HMI tags "MixingHead"
   "DB611_Hydraulic_State_Read" : Bool = PLC DB611_Hydraulic_State.Read AT %DB611.DBX8.0, 1 s
   "DB611_Hydraulic_State_Write" : Bool = PLC DB14_TP_Shortcuts.TP_Shortcuts.PageNo.7 AT %DB611.DBX8.1, 1 s
   "DB721_MH_Hydraulic_MH_Hyd{0}_Hyd_CP_Time" : S5Time = PLC DB14_TP_Shortcuts.TP_Shortcuts.PageNo.3 AT %DB721.DBW18, 1 s
      on ChangeValue: SetBit("DB611_Hydraulic_State_Write")
   "DB721_MH_Hydraulic_MH_Hyd{0}_Hyd_P_Startup" : S5Time = PLC DB14_TP_Shortcuts.TP_Shortcuts.PageNo.2 AT %DB721.DBW14, 1 s
      on ChangeValue: SetBit("DB611_Hydraulic_State_Write")
   "DB721_MH_Hydraulic_MH_Hyd{0}_Hyd_P_Supervision" : S5Time = PLC DB14_TP_Shortcuts.TP_Shortcuts.PageNo.4 AT %DB721.DBW16, 1 s
      on ChangeValue: SetBit("DB611_Hydraulic_State_Write")
   "DB721_MH_Hydraulic_MH_Hyd{0}_Hyd_PressureSwitch" : S5Time = PLC DB14_TP_Shortcuts.TP_Shortcuts.PageNo.5 AT %DB721.DBW20, 1 s
      on ChangeValue: SetBit("DB611_Hydraulic_State_Write")
   "DB721_MH_Hydraulic_MH_Hyd{0}_Hyd_SwitchOFFDelay" : S5Time = PLC DB14_TP_Shortcuts.TP_Shortcuts.PageNo.6 AT %DB721.DBW22, 1 s
      on ChangeValue: SetBit("DB611_Hydraulic_State_Write")
   "DB721_MH_Hydraulic_Option{0}_With2PSwitch" : Bool = PLC DB721_MH_Hydraulic.Option[0].With2PSwitch AT %DB721.DBX6.0, 1 s
   "MixingHead Options" : Int, internal
   "DB704_MH_Value_Read" : Bool = PLC DB704_MH_Value.Read AT %DB704.DBX4.0, 1 s
   "DB614_MH_State_Read" : Bool = PLC DB614_MH_State.Read AT %DB614.DBX8.0, 1 s
   "DB614_MH_State_Write" : Bool = PLC DB614_MH_State.Write AT %DB614.DBX8.1, 1 s
   "DB614_MH_State_MH_Status{0}_QPB_Values_selected" : Bool = PLC DB614_MH_State.MH_Status[0].QPB_Values_selected AT %DB614.DBX3920.2, 1 s
   "DB704_MH_Value_MH_Inerting{0}_Purge_time" : S5Time = PLC DB704_MH_Value.MH_Inerting[0].Purge_time AT %DB704.DBW4568, 1 s
      on ChangeValue: SetBit("DB704_MH_Value_Write")
   "DB704_MH_Value_MH_Inerting{0}_Purge_after_Shot" : S5Time = PLC DB704_MH_Value.MH_Inerting[0].Purge_after_Shot AT %DB704.DBW4570, 1 s
      on ChangeValue: SetBit("DB704_MH_Value_Write")
   "DB704_MH_Value_Mixinghead{0}_MH_Connection{1}_Flow_red_Circ" : Real = PLC DB704_MH_Value.Mixinghead[0].MH_Connection[1].Flow_red_Circ AT %DB704.DBD74, 1 s
      on ChangeValue: SetBit("DB704_MH_Value_Write")
   "DB704_MH_Value_Mixinghead{0}_MH_Connection{1}_Flow_HP_Circ" : Real = PLC DB704_MH_Value.Mixinghead[0].MH_Connection[1].Flow_HP_Circ AT %DB704.DBD70, 1 s
      on ChangeValue: SetBit("DB704_MH_Value_Write")
   "DB704_MH_Value_Mixinghead{0}_MH_Connection{1}_Flow_LP_Circ" : Real = PLC DB704_MH_Value.Mixinghead[0].MH_Connection[1].Flow_LP_Circ AT %DB704.DBD78, 1 s
      on ChangeValue: SetBit("DB704_MH_Value_Write")
   "DB704_MH_Value_Mixinghead{0}_MH_Connection{2}_Flow_HP_Circ" : Real = PLC DB704_MH_Value.Mixinghead[0].MH_Connection[2].Flow_HP_Circ AT %DB704.DBD104, 1 s
      on ChangeValue: SetBit("DB704_MH_Value_Write")
   "DB704_MH_Value_Mixinghead{0}_MH_Connection{2}_Flow_red_Circ" : Real = PLC DB704_MH_Value.Mixinghead[0].MH_Connection[2].Flow_red_Circ AT %DB704.DBD108, 1 s
      on ChangeValue: SetBit("DB704_MH_Value_Write")
   "DB704_MH_Value_Mixinghead{0}_MH_Connection{2}_Flow_LP_Circ" : Real = PLC DB704_MH_Value.Mixinghead[0].MH_Connection[2].Flow_LP_Circ AT %DB704.DBD112, 1 s
      on ChangeValue: SetBit("DB704_MH_Value_Write")
   "DB704_MH_Value_Mixinghead{0}_MH_Connection{1}_FlowQPB" : Real = PLC DB704_MH_Value.Mixinghead[0].MH_Connection[1].FlowQPB AT %DB704.DBD90, 1 s
      on ChangeValue: SetBit("DB704_MH_Value_Write")
   "DB704_MH_Value_Mixinghead{0}_MH_Connection{1}_HP_CircOverNozzle" : Bool = PLC DB704_MH_Value.Mixinghead[0].MH_Connection[1].HP_CircOverNozzle AT %DB704.DBX98.0, 1 s
      on ChangeValue: SetBit("DB614_MH_State_Write")
   "DB704_MH_Value_Mixinghead{0}_MH_Connection{1}_Red_CircOverNozzle" : Bool = PLC DB704_MH_Value.Mixinghead[0].MH_Connection[1].Red_CircOverNozzle AT %DB704.DBX98.1, 1 s
      on ChangeValue: SetBit("DB614_MH_State_Write")
   "DB704_MH_Value_Mixinghead{0}_MH_Connection{1}_LP_CircOverNozzle" : Bool = PLC DB704_MH_Value.Mixinghead[0].MH_Connection[1].LP_CircOverNozzle AT %DB704.DBX98.2, 1 s
      on ChangeValue: SetBit("DB614_MH_State_Write")
   "DB704_MH_Value_Mixinghead{0}_MH_Connection{2}_HP_CircOverNozzle" : Bool = PLC DB704_MH_Value.Mixinghead[0].MH_Connection[2].HP_CircOverNozzle AT %DB704.DBX132.0, 1 s
      on ChangeValue: SetBit("DB614_MH_State_Write")
   "DB704_MH_Value_Mixinghead{0}_MH_Connection{2}_Red_CircOverNozzle" : Bool = PLC DB704_MH_Value.Mixinghead[0].MH_Connection[2].Red_CircOverNozzle AT %DB704.DBX132.1, 1 s
      on ChangeValue: SetBit("DB614_MH_State_Write")
   "DB704_MH_Value_Mixinghead{0}_MH_Connection{2}_LP_CircOverNozzle" : Bool = PLC DB704_MH_Value.Mixinghead[0].MH_Connection[2].LP_CircOverNozzle AT %DB704.DBX132.2, 1 s
      on ChangeValue: SetBit("DB614_MH_State_Write")
   "MH_Control_Visibility" : Int AT %DB1.DBX0.0
   "DB704_MH_Value_Mixinghead{0}_MH_Connection{2}_FlowQPB" : Real = PLC DB704_MH_Value.Mixinghead[0].MH_Connection[2].FlowQPB AT %DB704.DBD124, 1 s
      on ChangeValue: SetBit("DB704_MH_Value_Write")
   "DB704_MH_Value_Mixinghead{0}_MH_Connection{2}_PressureQPB" : Real = PLC DB704_MH_Value.Mixinghead[0].MH_Connection[2].PressureQPB AT %DB704.DBD128, 1 s
      on ChangeValue: SetBit("DB704_MH_Value_Write")
   "DB704_MH_Value_Mixinghead{0}_MH_Connection{1}_PressureQPB" : Real = PLC DB704_MH_Value.Mixinghead[0].MH_Connection[1].PressureQPB AT %DB704.DBD94, 1 s
      on ChangeValue: SetBit("DB704_MH_Value_Write")
   "DB704_MH_Value_Mixinghead{0}_Cleaning_Piston_RestTimeBack" : S5Time = PLC DB704_MH_Value.Mixinghead[0].Cleaning_Piston.RestTimeBack AT %DB704.DBW44, 1 s
      on ChangeValue: SetBit("DB704_MH_Value_Write")
   "DB704_MH_Value_Mixinghead{0}_Cleaning_Piston_RestTimeFront" : S5Time = PLC DB704_MH_Value.Mixinghead[0].Cleaning_Piston.RestTimeFront AT %DB704.DBW46, 1 s
      on ChangeValue: SetBit("DB704_MH_Value_Write")
   "DB704_MH_Value_Mixinghead{0}_Cleaning_Piston_RestTimeFrontManual" : S5Time = PLC DB704_MH_Value.Mixinghead[0].Cleaning_Piston.RestTimeFrontManual AT %DB704.DBW48, 1 s
      on ChangeValue: SetBit("DB704_MH_Value_Write")
   "DB704_MH_Value_Write" : Bool = PLC DB704_MH_Value.Write AT %DB704.DBX4.1, 1 s
   "DB704_MH_Value_MH_Inerting{0}_Max_Inerting_Time" : S5Time = PLC DB704_MH_Value.MH_Inerting[0].Max_Inerting_Time AT %DB704.DBW4560, 1 s
      on ChangeValue: SetBit("DB704_MH_Value_Write")
   "DB704_MH_Value_MH_Inerting{0}_Ready_Time_after_Inert" : S5Time = PLC DB704_MH_Value.MH_Inerting[0].Ready_Time_after_Inert AT %DB704.DBW4562, 1 s
      on ChangeValue: SetBit("DB704_MH_Value_Write")
   "DB704_MH_Value_MH_Inerting{0}_Foam_density" : DInt = PLC DB704_MH_Value.MH_Inerting[0].Foam_density AT %DB704.DBD4538, 1 s
      on ChangeValue: SetBit("DB704_MH_Value_Write")
   "DB704_MH_Value_MH_Inerting{0}_Inerting_factor" : Real = PLC DB704_MH_Value.MH_Inerting[0].Inerting_factor AT %DB704.DBD4542, 1 s
      on ChangeValue: SetBit("DB704_MH_Value_Write")
   "DB704_MH_Value_MH_Inerting{0}_Start_Offset" : Real = PLC DB704_MH_Value.MH_Inerting[0].Start_Offset AT %DB704.DBD4546, 1 s
      on ChangeValue: SetBit("DB704_MH_Value_Write")
   "DB704_MH_Value_MH_Inerting{0}_Leakage_Value" : Real = PLC DB704_MH_Value.MH_Inerting[0].Leakage_Value AT %DB704.DBD4550, 1 s
      on ChangeValue: SetBit("DB704_MH_Value_Write")
   "DB704_MH_Value_Mixinghead{0}_AmountComponent" : Byte = PLC DB704_MH_Value.Mixinghead[0].AmountComponent AT %DB704.DBB6, 1 s
      on ChangeValue: SetBit("DB704_MH_Value_Write")
   "DB704_MH_Value_Mixinghead{0}_MachineNumber" : Byte = PLC DB704_MH_Value.Mixinghead[0].MachineNumber AT %DB704.DBB7, 1 s
      on ChangeValue: SetBit("DB704_MH_Value_Write")
   "DB704_MH_Value_Mixinghead{0}_MH_Active" : Bool = PLC DB704_MH_Value.Mixinghead[0].MH_Active AT %DB704.DBX9.0, 1 s
      on ChangeValue: SetBit("DB614_MH_State_Write")
   "DB704_MH_Value_Mixinghead{0}_With99program" : Bool = PLC DB704_MH_Value.Mixinghead[0].With99program AT %DB704.DBX10.2, 1 s
      on ChangeValue: SetBit("DB704_MH_Value_Write")
   "DB704_MH_Value_Mixinghead{0}_WithHeating" : Bool = PLC DB704_MH_Value.Mixinghead[0].WithHeating AT %DB704.DBX9.6, 1 s
      on ChangeValue: SetBit("DB704_MH_Value_Write")
   "DB704_MH_Value_Mixinghead{0}_WithInerting" : Bool = PLC DB704_MH_Value.Mixinghead[0].WithInerting AT %DB704.DBX9.5, 1 s
      on ChangeValue: SetBit("DB704_MH_Value_Write")
   "DB704_MH_Value_Mixinghead{0}_WithInterface" : Bool = PLC DB704_MH_Value.Mixinghead[0].WithInterface AT %DB704.DBX9.4, 1 s
      on ChangeValue: SetBit("DB704_MH_Value_Write")
   "DB704_MH_Value_Mixinghead{0}_WithNozzleControl" : Bool = PLC DB704_MH_Value.Mixinghead[0].WithNozzleControl AT %DB704.DBX9.2, 1 s
      on ChangeValue: SetBit("DB704_MH_Value_Write")
   "DB704_MH_Value_Mixinghead{0}_WithCleaningPiston" : Bool = PLC DB704_MH_Value.Mixinghead[0].WithCleaningPiston AT %DB704.DBX9.1, 1 s
      on ChangeValue: SetBit("DB704_MH_Value_Write")
   "DB704_MH_Value_Mixinghead{0}_WithLPCirculation" : Bool = PLC DB704_MH_Value.Mixinghead[0].WithLPCirculation AT %DB704.DBX9.3, 1 s
      on ChangeValue: SetBit("DB704_MH_Value_Write")
   "DB704_MH_Value_Mixinghead{0}_pRrgNumberManual" : Byte = PLC DB704_MH_Value.Mixinghead[0].pRrgNumberManual AT %DB704.DBB8, 1 s
      on ChangeValue: SetBit("DB704_MH_Value_Write")
   "DB704_MH_Value_Mixinghead{0}_Openingtime" : Real = PLC DB704_MH_Value.Mixinghead[0].Openingtime AT %DB704.DBD14, 1 s
      on ChangeValue: SetBit("DB704_MH_Value_Write")
   "DB704_MH_Value_Mixinghead{0}_Closingtime" : Real = PLC DB704_MH_Value.Mixinghead[0].Closingtime AT %DB704.DBD18, 1 s
      on ChangeValue: SetBit("DB704_MH_Value_Write")
   "DB604_PV_Mixinghead_Mixinghead{0}_Temperature_Connection{1}_PV_ActV_Value" : Real = PLC DB604_PV_Mixinghead.Mixinghead[0].Temperature_Connection[1].PV_ActV.Value AT %DB604.DBD314, 1 s
      on ChangeValue: SetBit("DB704_MH_Value_Write")
   "DB604_PV_Mixinghead_Mixinghead{0}_Temperature_Connection{1}_PV_SetV_Value" : Real = PLC DB604_PV_Mixinghead.Mixinghead[0].Temperature_Connection[1].PV_SetV.Value AT %DB604.DBD294, 1 s
      on ChangeValue: SetBit("DB704_MH_Value_Write")
   "DB604_PV_Mixinghead_Mixinghead{0}_Temperature_Connection{1}_PV_SetV_WarningLowerLimit" : Real = PLC DB604_PV_Mixinghead.Mixinghead[0].Temperature_Connection[1].PV_SetV.WarningLowerLimit AT %DB604.DBD298, 1 s
      on ChangeValue: SetBit("DB704_MH_Value_Write")
   "DB604_PV_Mixinghead_Mixinghead{0}_Temperature_Connection{1}_PV_SetV_WarningUpperLimit" : Real = PLC DB604_PV_Mixinghead.Mixinghead[0].Temperature_Connection[1].PV_SetV.WarningUpperLimit AT %DB604.DBD302, 1 s
      on ChangeValue: SetBit("DB704_MH_Value_Write")
   "DB604_PV_Mixinghead_Mixinghead{0}_Temperature_Connection{1}_PV_SetV_AlarmLowerLimit" : Real = PLC DB604_PV_Mixinghead.Mixinghead[0].Temperature_Connection[1].PV_SetV.AlarmLowerLimit AT %DB604.DBD306, 1 s
      on ChangeValue: SetBit("DB704_MH_Value_Write")
   "DB604_PV_Mixinghead_Mixinghead{0}_Temperature_Connection{1}_PV_SetV_AlarmUpperLimit" : Real = PLC DB604_PV_Mixinghead.Mixinghead[0].Temperature_Connection[1].PV_SetV.AlarmUpperLimit AT %DB604.DBD310, 1 s
      on ChangeValue: SetBit("DB704_MH_Value_Write")
   "DB604_PV_Mixinghead_Mixinghead{0}_Pressure_Connection{1}_PV_SetV_Value" : Real = PLC DB604_PV_Mixinghead.Mixinghead[0].Pressure_Connection[1].PV_SetV.Value AT %DB604.DBD6, 1 s
      on ChangeValue: SetBit("DB704_MH_Value_Write")
   "DB604_PV_Mixinghead_Mixinghead{0}_Pressure_Connection{1}_PV_SetV_WarningLowerLimit" : Real = PLC DB604_PV_Mixinghead.Mixinghead[0].Pressure_Connection[1].PV_SetV.WarningLowerLimit AT %DB604.DBD10, 1 s
      on ChangeValue: SetBit("DB704_MH_Value_Write")
   "DB604_PV_Mixinghead_Mixinghead{0}_Pressure_Connection{1}_PV_SetV_WarningUpperLimit" : Real = PLC DB604_PV_Mixinghead.Mixinghead[0].Pressure_Connection[1].PV_SetV.WarningUpperLimit AT %DB604.DBD14, 1 s
      on ChangeValue: SetBit("DB704_MH_Value_Write")
   "DB604_PV_Mixinghead_Mixinghead{0}_Pressure_Connection{1}_PV_SetV_AlarmLowerLimit" : Real = PLC DB604_PV_Mixinghead.Mixinghead[0].Pressure_Connection[1].PV_SetV.AlarmLowerLimit AT %DB604.DBD18, 1 s
      on ChangeValue: SetBit("DB704_MH_Value_Write")
   "DB604_PV_Mixinghead_Mixinghead{0}_Pressure_Connection{1}_PV_SetV_AlarmUpperLimit" : Real = PLC DB604_PV_Mixinghead.Mixinghead[0].Pressure_Connection[1].PV_SetV.AlarmUpperLimit AT %DB604.DBD22, 1 s
      on ChangeValue: SetBit("DB704_MH_Value_Write")
   "DB604_PV_Mixinghead_Mixinghead{0}_Pressure_Connection{1}_PV_ActV_Value" : Real = PLC DB604_PV_Mixinghead.Mixinghead[0].Pressure_Connection[1].PV_ActV.Value AT %DB604.DBD26, 1 s
      on ChangeValue: SetBit("DB704_MH_Value_Write")
   "DB604_PV_Mixinghead_Mixinghead{0}_Pressure_Connection{2}_PV_SetV_Value" : Real = PLC DB604_PV_Mixinghead.Mixinghead[0].Pressure_Connection[2].PV_SetV.Value AT %DB604.DBD54, 1 s
      on ChangeValue: SetBit("DB704_MH_Value_Write")
   "DB604_PV_Mixinghead_Mixinghead{0}_Pressure_Connection{2}_PV_SetV_WarningLowerLimit" : Real = PLC DB604_PV_Mixinghead.Mixinghead[0].Pressure_Connection[2].PV_SetV.WarningLowerLimit AT %DB604.DBD58, 1 s
      on ChangeValue: SetBit("DB704_MH_Value_Write")
   "DB604_PV_Mixinghead_Mixinghead{0}_Pressure_Connection{2}_PV_SetV_WarningUpperLimit" : Real = PLC DB604_PV_Mixinghead.Mixinghead[0].Pressure_Connection[2].PV_SetV.WarningUpperLimit AT %DB604.DBD62, 1 s
      on ChangeValue: SetBit("DB704_MH_Value_Write")
   "DB604_PV_Mixinghead_Mixinghead{0}_Pressure_Connection{2}_PV_SetV_AlarmLowerLimit" : Real = PLC DB604_PV_Mixinghead.Mixinghead[0].Pressure_Connection[2].PV_SetV.AlarmLowerLimit AT %DB604.DBD66, 1 s
      on ChangeValue: SetBit("DB704_MH_Value_Write")
   "DB604_PV_Mixinghead_Mixinghead{0}_Pressure_Connection{2}_PV_SetV_AlarmUpperLimit" : Real = PLC DB604_PV_Mixinghead.Mixinghead[0].Pressure_Connection[2].PV_SetV.AlarmUpperLimit AT %DB604.DBD70, 1 s
      on ChangeValue: SetBit("DB704_MH_Value_Write")
   "DB604_PV_Mixinghead_Mixinghead{0}_Pressure_Connection{2}_PV_ActV_Value" : Real = PLC DB604_PV_Mixinghead.Mixinghead[0].Pressure_Connection[2].PV_ActV.Value AT %DB604.DBD74, 1 s
      on ChangeValue: SetBit("DB704_MH_Value_Write")
   "DB604_PV_Mixinghead_Mixinghead{0}_Temperature_Connection{2}_PV_SetV_Value" : Real = PLC DB604_PV_Mixinghead.Mixinghead[0].Temperature_Connection[2].PV_SetV.Value AT %DB604.DBD342, 1 s
      on ChangeValue: SetBit("DB704_MH_Value_Write")
   "DB604_PV_Mixinghead_Mixinghead{0}_Temperature_Connection{2}_PV_SetV_WarningLowerLimit" : Real = PLC DB604_PV_Mixinghead.Mixinghead[0].Temperature_Connection[2].PV_SetV.WarningLowerLimit AT %DB604.DBD346, 1 s
      on ChangeValue: SetBit("DB704_MH_Value_Write")
   "DB604_PV_Mixinghead_Mixinghead{0}_Temperature_Connection{2}_PV_SetV_WarningUpperLimit" : Real = PLC DB604_PV_Mixinghead.Mixinghead[0].Temperature_Connection[2].PV_SetV.WarningUpperLimit AT %DB604.DBD350, 1 s
      on ChangeValue: SetBit("DB704_MH_Value_Write")
   "DB604_PV_Mixinghead_Mixinghead{0}_Temperature_Connection{2}_PV_SetV_AlarmLowerLimit" : Real = PLC DB604_PV_Mixinghead.Mixinghead[0].Temperature_Connection[2].PV_SetV.AlarmLowerLimit AT %DB604.DBD354, 1 s
      on ChangeValue: SetBit("DB704_MH_Value_Write")
   "DB604_PV_Mixinghead_Mixinghead{0}_Temperature_Connection{2}_PV_SetV_AlarmUpperLimit" : Real = PLC DB604_PV_Mixinghead.Mixinghead[0].Temperature_Connection[2].PV_SetV.AlarmUpperLimit AT %DB604.DBD358, 1 s
      on ChangeValue: SetBit("DB704_MH_Value_Write")
   "DB604_PV_Mixinghead_Mixinghead{0}_Temperature_Connection{2}_PV_ActV_Value" : Real = PLC DB604_PV_Mixinghead.Mixinghead[0].Temperature_Connection[2].PV_ActV.Value AT %DB604.DBD362, 1 s
      on ChangeValue: SetBit("DB704_MH_Value_Write")
   "DB704_MH_Value_Mixinghead{0}_Cleaning_Piston_CP_withInterval" : Bool = PLC DB704_MH_Value.Mixinghead[0].Cleaning_Piston.CP_withInterval AT %DB704.DBX56.1, 1 s
      on ChangeValue: SetBit("DB704_MH_Value_Write")
   "DB704_MH_Value_Mixinghead{0}_Cleaning_Piston_ContrCleaningPiston" : Bool = PLC DB704_MH_Value.Mixinghead[0].Cleaning_Piston.ContrCleaningPiston AT %DB704.DBX56.3, 1 s
      on ChangeValue: SetBit("DB704_MH_Value_Write")
   "DB611_Hydraulic_State_MH_Hydraulic{0}_HourCounter" : DInt = PLC DB611_Hydraulic_State.MH_Hydraulic[0].HourCounter AT %DB611.DBD14, 1 s
   "DB614_MH_State_ReadDeviceNo" : Int = PLC DB614_MH_State.ReadDeviceNo AT %DB614.DBW0, 1 s
   "DB704_MH_Value_Mixinghead{0}_WithMHVenting" : Bool = PLC DB704_MH_Value.Mixinghead[0].WithMHVenting AT %DB704.DBX9.7, 1 s
      on ChangeValue: SetBit("DB704_MH_Value_Write")
   "DB614_MH_State_MH_Status{0}_Switch_HP_ON_OFF" : Bool = PLC DB614_MH_State.MH_Status[0].Switch_HP_ON_OFF AT %DB614.DBX3920.5, 1 s
      on ChangeValue: SetBit("DB614_MH_State_Write")
   "DB614_MH_State_MH_Status{0}_Switch_Service_ON_OFF" : Bool = PLC DB614_MH_State.MH_Status[0].Switch_Service_ON_OFF AT %DB614.DBX3920.6, 1 s
      on ChangeValue: SetBit("DB614_MH_State_Write")
   "DB704_MH_Value_Mixinghead{0}_MH_Connection{3}_Flow_HP_Circ" : Real = PLC DB704_MH_Value.Mixinghead[0].MH_Connection[3].Flow_HP_Circ AT %DB704.DBD138, 1 s
   "DB704_MH_Value_Mixinghead{0}_MH_Connection{3}_Flow_red_Circ" : Real = PLC DB704_MH_Value.Mixinghead[0].MH_Connection[3].Flow_red_Circ AT %DB704.DBD142, 1 s
   "DB704_MH_Value_Mixinghead{0}_MH_Connection{3}_Flow_LP_Circ" : Real = PLC DB704_MH_Value.Mixinghead[0].MH_Connection[3].Flow_LP_Circ AT %DB704.DBD146, 1 s
   "DB704_MH_Value_Mixinghead{0}_MH_Connection{3}_HP_CircOverNozzle" : Bool = PLC DB704_MH_Value.Mixinghead[0].MH_Connection[3].HP_CircOverNozzle AT %DB704.DBX166.0, 1 s
   "DB704_MH_Value_Mixinghead{0}_MH_Connection{3}_Red_CircOverNozzle" : Bool = PLC DB704_MH_Value.Mixinghead[0].MH_Connection[3].Red_CircOverNozzle AT %DB704.DBX166.1, 1 s
   "DB704_MH_Value_Mixinghead{0}_MH_Connection{3}_LP_CircOverNozzle" : Bool = PLC DB704_MH_Value.Mixinghead[0].MH_Connection[3].LP_CircOverNozzle AT %DB704.DBX166.2, 1 s
   "DB704_MH_Value_Mixinghead{0}_MH_Connection{4}_Flow_HP_Circ" : Real = PLC DB704_MH_Value.Mixinghead[0].MH_Connection[4].Flow_HP_Circ AT %DB704.DBD172, 1 s
   "DB704_MH_Value_Mixinghead{0}_MH_Connection{4}_Flow_red_Circ" : Real = PLC DB704_MH_Value.Mixinghead[0].MH_Connection[4].Flow_red_Circ AT %DB704.DBD176, 1 s
   "DB704_MH_Value_Mixinghead{0}_MH_Connection{4}_Flow_LP_Circ" : Real = PLC DB704_MH_Value.Mixinghead[0].MH_Connection[4].Flow_LP_Circ AT %DB704.DBD180, 1 s
   "DB704_MH_Value_Mixinghead{0}_MH_Connection{4}_HP_CircOverNozzle" : Bool = PLC DB704_MH_Value.Mixinghead[0].MH_Connection[4].HP_CircOverNozzle AT %DB704.DBX200.0, 1 s
   "DB704_MH_Value_Mixinghead{0}_MH_Connection{4}_Red_CircOverNozzle" : Bool = PLC DB702_Tank_Value.Tank[0].With_Drain AT %DB704.DBX200.1, 1 s
   "DB704_MH_Value_Mixinghead{0}_MH_Connection{4}_LP_CircOverNozzle" : Bool = PLC DB704_MH_Value.Mixinghead[0].MH_Connection[4].LP_CircOverNozzle AT %DB704.DBX200.2, 1 s
   "DB704_MH_Value_Mixinghead{0}_MH_Connection{5}_Flow_HP_Circ" : Real = PLC DB704_MH_Value.Mixinghead[0].MH_Connection[5].Flow_HP_Circ AT %DB704.DBD206, 1 s
   "DB704_MH_Value_Mixinghead{0}_MH_Connection{5}_Flow_red_Circ" : Real = PLC DB704_MH_Value.Mixinghead[0].MH_Connection[5].Flow_red_Circ AT %DB704.DBD210, 1 s
   "DB704_MH_Value_Mixinghead{0}_MH_Connection{5}_Flow_LP_Circ" : Real = PLC DB704_MH_Value.Mixinghead[0].MH_Connection[5].Flow_LP_Circ AT %DB704.DBD214, 1 s
   "DB704_MH_Value_Mixinghead{0}_MH_Connection{5}_HP_CircOverNozzle" : Bool = PLC DB704_MH_Value.Mixinghead[0].MH_Connection[5].HP_CircOverNozzle AT %DB704.DBX234.0, 1 s
   "DB704_MH_Value_Mixinghead{0}_MH_Connection{5}_Red_CircOverNozzle" : Bool = PLC DB704_MH_Value.Mixinghead[0].MH_Connection[5].Red_CircOverNozzle AT %DB704.DBX234.1, 1 s
   "DB704_MH_Value_Mixinghead{0}_MH_Connection{5}_LP_CircOverNozzle" : Bool = PLC DB704_MH_Value.Mixinghead[0].MH_Connection[5].LP_CircOverNozzle AT %DB704.DBX234.2, 1 s
   "DB704_MH_Value_Mixinghead{0}_MH_Connection{6}_Flow_HP_Circ" : Real = PLC DB704_MH_Value.Mixinghead[0].MH_Connection[6].Flow_HP_Circ AT %DB704.DBD240, 1 s
   "DB704_MH_Value_Mixinghead{0}_MH_Connection{6}_Flow_red_Circ" : Real = PLC DB704_MH_Value.Mixinghead[0].MH_Connection[6].Flow_red_Circ AT %DB704.DBD244, 1 s
   "DB704_MH_Value_Mixinghead{0}_MH_Connection{6}_Flow_LP_Circ" : Real = PLC DB704_MH_Value.Mixinghead[0].MH_Connection[6].Flow_LP_Circ AT %DB704.DBD248, 1 s
   "DB704_MH_Value_Mixinghead{0}_MH_Connection{6}_HP_CircOverNozzle" : Bool = PLC DB704_MH_Value.Mixinghead[0].MH_Connection[6].HP_CircOverNozzle AT %DB704.DBX268.0, 1 s
   "DB704_MH_Value_Mixinghead{0}_MH_Connection{6}_Red_CircOverNozzle" : Bool = PLC DB704_MH_Value.Mixinghead[0].MH_Connection[6].Red_CircOverNozzle AT %DB704.DBX268.1, 1 s
   "DB704_MH_Value_Mixinghead{0}_MH_Connection{6}_LP_CircOverNozzle" : Bool = PLC DB704_MH_Value.Mixinghead[0].MH_Connection[6].LP_CircOverNozzle AT %DB704.DBX268.2, 1 s
   "DB704_MH_Value_Mixinghead{0}_MH_Connection{3}_FlowQPB" : Real = PLC DB704_MH_Value.Mixinghead[0].MH_Connection[3].FlowQPB AT %DB704.DBD158, 1 s
   "DB704_MH_Value_Mixinghead{0}_MH_Connection{3}_PressureQPB" : Real = PLC DB704_MH_Value.Mixinghead[0].MH_Connection[3].PressureQPB AT %DB704.DBD162, 1 s
   "DB704_MH_Value_Mixinghead{0}_MH_Connection{4}_FlowQPB" : Real = PLC DB704_MH_Value.Mixinghead[0].MH_Connection[4].FlowQPB AT %DB704.DBD192, 1 s
   "DB704_MH_Value_Mixinghead{0}_MH_Connection{4}_PressureQPB" : Real = PLC DB704_MH_Value.Mixinghead[0].MH_Connection[4].PressureQPB AT %DB704.DBD196, 1 s
   "DB704_MH_Value_Mixinghead{0}_MH_Connection{5}_FlowQPB" : Real = PLC DB704_MH_Value.Mixinghead[0].MH_Connection[5].FlowQPB AT %DB704.DBD226, 1 s
   "DB704_MH_Value_Mixinghead{0}_MH_Connection{5}_PressureQPB" : Real = PLC DB704_MH_Value.Mixinghead[0].MH_Connection[5].PressureQPB AT %DB704.DBD230, 1 s
   "DB704_MH_Value_Mixinghead{0}_MH_Connection{6}_FlowQPB" : Real = PLC DB704_MH_Value.Mixinghead[0].MH_Connection[6].FlowQPB AT %DB704.DBD260, 1 s
   "DB704_MH_Value_Mixinghead{0}_MH_Connection{6}_PressureQPB" : Real = PLC DB704_MH_Value.Mixinghead[0].MH_Connection[6].PressureQPB AT %DB704.DBD264, 1 s
   "DB604_PV_Mixinghead_Mixinghead{0}_Temperature_Connection{3}_PV_ActV_Value" : Real = PLC DB604_PV_Mixinghead.Mixinghead[0].Temperature_Connection[3].PV_ActV.Value AT %DB604.DBD410, 1 s
      on ChangeValue: SetBit("DB704_MH_Value_Write")
   "DB604_PV_Mixinghead_Mixinghead{0}_Temperature_Connection{3}_PV_SetV_Value" : Real = PLC DB604_PV_Mixinghead.Mixinghead[0].Temperature_Connection[3].PV_SetV.Value AT %DB604.DBD390, 1 s
      on ChangeValue: SetBit("DB704_MH_Value_Write")
   "DB604_PV_Mixinghead_Mixinghead{0}_Temperature_Connection{3}_PV_SetV_WarningLowerLimit" : Real = PLC DB604_PV_Mixinghead.Mixinghead[0].Temperature_Connection[3].PV_SetV.WarningLowerLimit AT %DB604.DBD394, 1 s
      on ChangeValue: SetBit("DB704_MH_Value_Write")
   "DB604_PV_Mixinghead_Mixinghead{0}_Temperature_Connection{3}_PV_SetV_WarningUpperLimit" : Real = PLC DB604_PV_Mixinghead.Mixinghead[0].Temperature_Connection[3].PV_SetV.WarningUpperLimit AT %DB604.DBD398, 1 s
      on ChangeValue: SetBit("DB704_MH_Value_Write")
   "DB604_PV_Mixinghead_Mixinghead{0}_Temperature_Connection{3}_PV_SetV_AlarmLowerLimit" : Real = PLC DB604_PV_Mixinghead.Mixinghead[0].Temperature_Connection[3].PV_SetV.AlarmLowerLimit AT %DB604.DBD402, 1 s
      on ChangeValue: SetBit("DB704_MH_Value_Write")
   "DB604_PV_Mixinghead_Mixinghead{0}_Temperature_Connection{3}_PV_SetV_AlarmUpperLimit" : Real = PLC DB604_PV_Mixinghead.Mixinghead[0].Temperature_Connection[3].PV_SetV.AlarmUpperLimit AT %DB604.DBD406, 1 s
      on ChangeValue: SetBit("DB704_MH_Value_Write")
   "DB604_PV_Mixinghead_Mixinghead{0}_Temperature_Connection{4}_PV_SetV_Value" : Real = PLC DB604_PV_Mixinghead.Mixinghead[0].Temperature_Connection[4].PV_SetV.Value AT %DB604.DBD438, 1 s
      on ChangeValue: SetBit("DB704_MH_Value_Write")
   "DB604_PV_Mixinghead_Mixinghead{0}_Temperature_Connection{4}_PV_SetV_WarningLowerLimit" : Real = PLC DB604_PV_Mixinghead.Mixinghead[0].Temperature_Connection[4].PV_SetV.WarningLowerLimit AT %DB604.DBD442, 1 s
      on ChangeValue: SetBit("DB704_MH_Value_Write")
   "DB604_PV_Mixinghead_Mixinghead{0}_Temperature_Connection{4}_PV_SetV_WarningUpperLimit" : Real = PLC DB604_PV_Mixinghead.Mixinghead[0].Temperature_Connection[4].PV_SetV.WarningUpperLimit AT %DB604.DBD446, 1 s
      on ChangeValue: SetBit("DB704_MH_Value_Write")
   "DB604_PV_Mixinghead_Mixinghead{0}_Temperature_Connection{4}_PV_SetV_AlarmLowerLimit" : Real = PLC DB604_PV_Mixinghead.Mixinghead[0].Temperature_Connection[4].PV_SetV.AlarmLowerLimit AT %DB604.DBD450, 1 s
      on ChangeValue: SetBit("DB704_MH_Value_Write")
   "DB604_PV_Mixinghead_Mixinghead{0}_Temperature_Connection{4}_PV_SetV_AlarmUpperLimit" : Real = PLC DB604_PV_Mixinghead.Mixinghead[0].Temperature_Connection[4].PV_SetV.AlarmUpperLimit AT %DB604.DBD454, 1 s
      on ChangeValue: SetBit("DB704_MH_Value_Write")
   "DB604_PV_Mixinghead_Mixinghead{0}_Temperature_Connection{4}_PV_ActV_Value" : Real = PLC DB604_PV_Mixinghead.Mixinghead[0].Temperature_Connection[4].PV_ActV.Value AT %DB604.DBD458, 1 s
      on ChangeValue: SetBit("DB704_MH_Value_Write")
   "DB604_PV_Mixinghead_Mixinghead{0}_Temperature_Connection{5}_PV_SetV_Value" : Real = PLC DB604_PV_Mixinghead.Mixinghead[0].Temperature_Connection[5].PV_SetV.Value AT %DB604.DBD486, 1 s
      on ChangeValue: SetBit("DB704_MH_Value_Write")
   "DB604_PV_Mixinghead_Mixinghead{0}_Temperature_Connection{5}_PV_SetV_WarningLowerLimit" : Real = PLC DB604_PV_Mixinghead.Mixinghead[0].Temperature_Connection[5].PV_SetV.WarningLowerLimit AT %DB604.DBD490, 1 s
      on ChangeValue: SetBit("DB704_MH_Value_Write")
   "DB604_PV_Mixinghead_Mixinghead{0}_Temperature_Connection{5}_PV_SetV_WarningUpperLimit" : Real = PLC DB604_PV_Mixinghead.Mixinghead[0].Temperature_Connection[5].PV_SetV.WarningUpperLimit AT %DB604.DBD494, 1 s
      on ChangeValue: SetBit("DB704_MH_Value_Write")
   "DB604_PV_Mixinghead_Mixinghead{0}_Temperature_Connection{5}_PV_SetV_AlarmLowerLimit" : Real = PLC DB604_PV_Mixinghead.Mixinghead[0].Temperature_Connection[5].PV_SetV.AlarmLowerLimit AT %DB604.DBD498, 1 s
      on ChangeValue: SetBit("DB704_MH_Value_Write")
   "DB604_PV_Mixinghead_Mixinghead{0}_Temperature_Connection{5}_PV_SetV_AlarmUpperLimit" : Real = PLC DB604_PV_Mixinghead.Mixinghead[0].Temperature_Connection[5].PV_SetV.AlarmUpperLimit AT %DB604.DBD502, 1 s
      on ChangeValue: SetBit("DB704_MH_Value_Write")
   "DB604_PV_Mixinghead_Mixinghead{0}_Temperature_Connection{5}_PV_ActV_Value" : Real = PLC DB604_PV_Mixinghead.Mixinghead[0].Temperature_Connection[5].PV_ActV.Value AT %DB604.DBD506, 1 s
      on ChangeValue: SetBit("DB704_MH_Value_Write")
   "DB604_PV_Mixinghead_Mixinghead{0}_Temperature_Connection{6}_PV_SetV_Value" : Real = PLC DB604_PV_Mixinghead.Mixinghead[0].Temperature_Connection[6].PV_SetV.Value AT %DB604.DBD534, 1 s
      on ChangeValue: SetBit("DB704_MH_Value_Write")
   "DB604_PV_Mixinghead_Mixinghead{0}_Temperature_Connection{6}_PV_SetV_WarningLowerLimit" : Real = PLC DB604_PV_Mixinghead.Mixinghead[0].Temperature_Connection[6].PV_SetV.WarningLowerLimit AT %DB604.DBD538, 1 s
      on ChangeValue: SetBit("DB704_MH_Value_Write")
   "DB604_PV_Mixinghead_Mixinghead{0}_Temperature_Connection{6}_PV_SetV_WarningUpperLimit" : Real = PLC DB604_PV_Mixinghead.Mixinghead[0].Temperature_Connection[6].PV_SetV.WarningUpperLimit AT %DB604.DBD542, 1 s
      on ChangeValue: SetBit("DB704_MH_Value_Write")
   "DB604_PV_Mixinghead_Mixinghead{0}_Temperature_Connection{6}_PV_SetV_AlarmLowerLimit" : Real = PLC DB604_PV_Mixinghead.Mixinghead[0].Temperature_Connection[6].PV_SetV.AlarmLowerLimit AT %DB604.DBD546, 1 s
      on ChangeValue: SetBit("DB704_MH_Value_Write")
   "DB604_PV_Mixinghead_Mixinghead{0}_Temperature_Connection{6}_PV_SetV_AlarmUpperLimit" : Real = PLC DB604_PV_Mixinghead.Mixinghead[0].Temperature_Connection[6].PV_SetV.AlarmUpperLimit AT %DB604.DBD550, 1 s
      on ChangeValue: SetBit("DB704_MH_Value_Write")
   "DB604_PV_Mixinghead_Mixinghead{0}_Temperature_Connection{6}_PV_ActV_Value" : Real = PLC DB604_PV_Mixinghead.Mixinghead[0].Temperature_Connection[6].PV_ActV.Value AT %DB604.DBD554, 1 s
      on ChangeValue: SetBit("DB704_MH_Value_Write")
   "DB604_PV_Mixinghead_Mixinghead{0}_Pressure_Connection{3}_PV_SetV_Value" : Real = PLC DB604_PV_Mixinghead.Mixinghead[0].Pressure_Connection[3].PV_SetV.Value AT %DB604.DBD102, 1 s
      on ChangeValue: SetBit("DB704_MH_Value_Write")
   "DB604_PV_Mixinghead_Mixinghead{0}_Pressure_Connection{3}_PV_SetV_WarningLowerLimit" : Real = PLC DB604_PV_Mixinghead.Mixinghead[0].Pressure_Connection[3].PV_SetV.WarningLowerLimit AT %DB604.DBD106, 1 s
      on ChangeValue: SetBit("DB704_MH_Value_Write")
   "DB604_PV_Mixinghead_Mixinghead{0}_Pressure_Connection{3}_PV_SetV_WarningUpperLimit" : Real = PLC DB604_PV_Mixinghead.Mixinghead[0].Pressure_Connection[3].PV_SetV.WarningUpperLimit AT %DB604.DBD110, 1 s
      on ChangeValue: SetBit("DB704_MH_Value_Write")
   "DB604_PV_Mixinghead_Mixinghead{0}_Pressure_Connection{3}_PV_SetV_AlarmLowerLimit" : Real = PLC DB604_PV_Mixinghead.Mixinghead[0].Pressure_Connection[3].PV_SetV.AlarmLowerLimit AT %DB604.DBD114, 1 s
      on ChangeValue: SetBit("DB704_MH_Value_Write")
   "DB604_PV_Mixinghead_Mixinghead{0}_Pressure_Connection{3}_PV_SetV_AlarmUpperLimit" : Real = PLC DB604_PV_Mixinghead.Mixinghead[0].Pressure_Connection[3].PV_SetV.AlarmUpperLimit AT %DB604.DBD118, 1 s
      on ChangeValue: SetBit("DB704_MH_Value_Write")
   "DB604_PV_Mixinghead_Mixinghead{0}_Pressure_Connection{3}_PV_ActV_Value" : Real = PLC DB604_PV_Mixinghead.Mixinghead[0].Pressure_Connection[3].PV_ActV.Value AT %DB604.DBD122, 1 s
      on ChangeValue: SetBit("DB704_MH_Value_Write")
   "DB604_PV_Mixinghead_Mixinghead{0}_Pressure_Connection{4}_PV_SetV_Value" : Real = PLC DB604_PV_Mixinghead.Mixinghead[0].Pressure_Connection[4].PV_SetV.Value AT %DB604.DBD150, 1 s
      on ChangeValue: SetBit("DB704_MH_Value_Write")
   "DB604_PV_Mixinghead_Mixinghead{0}_Pressure_Connection{4}_PV_SetV_WarningLowerLimit" : Real = PLC DB604_PV_Mixinghead.Mixinghead[0].Pressure_Connection[4].PV_SetV.WarningLowerLimit AT %DB604.DBD154, 1 s
      on ChangeValue: SetBit("DB704_MH_Value_Write")
   "DB604_PV_Mixinghead_Mixinghead{0}_Pressure_Connection{4}_PV_SetV_WarningUpperLimit" : Real = PLC DB604_PV_Mixinghead.Mixinghead[0].Pressure_Connection[4].PV_SetV.WarningUpperLimit AT %DB604.DBD158, 1 s
      on ChangeValue: SetBit("DB704_MH_Value_Write")
   "DB604_PV_Mixinghead_Mixinghead{0}_Pressure_Connection{4}_PV_SetV_AlarmLowerLimit" : Real = PLC DB604_PV_Mixinghead.Mixinghead[0].Pressure_Connection[4].PV_SetV.AlarmLowerLimit AT %DB604.DBD162, 1 s
      on ChangeValue: SetBit("DB704_MH_Value_Write")
   "DB604_PV_Mixinghead_Mixinghead{0}_Pressure_Connection{4}_PV_SetV_AlarmUpperLimit" : Real = PLC DB604_PV_Mixinghead.Mixinghead[0].Pressure_Connection[4].PV_SetV.AlarmUpperLimit AT %DB604.DBD166, 1 s
      on ChangeValue: SetBit("DB704_MH_Value_Write")
   "DB604_PV_Mixinghead_Mixinghead{0}_Pressure_Connection{4}_PV_ActV_Value" : Real = PLC DB604_PV_Mixinghead.Mixinghead[0].Pressure_Connection[4].PV_ActV.Value AT %DB604.DBD170, 1 s
      on ChangeValue: SetBit("DB704_MH_Value_Write")
   "DB604_PV_Mixinghead_Mixinghead{0}_Pressure_Connection{5}_PV_SetV_Value" : Real = PLC DB604_PV_Mixinghead.Mixinghead[0].Pressure_Connection[5].PV_SetV.Value AT %DB604.DBD198, 1 s
      on ChangeValue: SetBit("DB704_MH_Value_Write")
   "DB604_PV_Mixinghead_Mixinghead{0}_Pressure_Connection{5}_PV_SetV_WarningLowerLimit" : Real = PLC DB604_PV_Mixinghead.Mixinghead[0].Pressure_Connection[5].PV_SetV.WarningLowerLimit AT %DB604.DBD202, 1 s
      on ChangeValue: SetBit("DB704_MH_Value_Write")
   "DB604_PV_Mixinghead_Mixinghead{0}_Pressure_Connection{5}_PV_SetV_WarningUpperLimit" : Real = PLC DB604_PV_Mixinghead.Mixinghead[0].Pressure_Connection[5].PV_SetV.WarningUpperLimit AT %DB604.DBD206, 1 s
      on ChangeValue: SetBit("DB704_MH_Value_Write")
   "DB604_PV_Mixinghead_Mixinghead{0}_Pressure_Connection{5}_PV_SetV_AlarmLowerLimit" : Real = PLC DB604_PV_Mixinghead.Mixinghead[0].Pressure_Connection[5].PV_SetV.AlarmLowerLimit AT %DB604.DBD210, 1 s
      on ChangeValue: SetBit("DB704_MH_Value_Write")
   "DB604_PV_Mixinghead_Mixinghead{0}_Pressure_Connection{5}_PV_SetV_AlarmUpperLimit" : Real = PLC DB604_PV_Mixinghead.Mixinghead[0].Pressure_Connection[5].PV_SetV.AlarmUpperLimit AT %DB604.DBD214, 1 s
      on ChangeValue: SetBit("DB704_MH_Value_Write")
   "DB604_PV_Mixinghead_Mixinghead{0}_Pressure_Connection{5}_PV_ActV_Value" : Real = PLC DB604_PV_Mixinghead.Mixinghead[0].Pressure_Connection[5].PV_ActV.Value AT %DB604.DBD218, 1 s
      on ChangeValue: SetBit("DB704_MH_Value_Write")
   "DB604_PV_Mixinghead_Mixinghead{0}_Pressure_Connection{6}_PV_SetV_Value" : Real = PLC DB604_PV_Mixinghead.Mixinghead[0].Pressure_Connection[6].PV_SetV.Value AT %DB604.DBD246, 1 s
      on ChangeValue: SetBit("DB704_MH_Value_Write")
   "DB604_PV_Mixinghead_Mixinghead{0}_Pressure_Connection{6}_PV_SetV_WarningLowerLimit" : Real = PLC DB604_PV_Mixinghead.Mixinghead[0].Pressure_Connection[6].PV_SetV.WarningLowerLimit AT %DB604.DBD250, 1 s
      on ChangeValue: SetBit("DB704_MH_Value_Write")
   "DB604_PV_Mixinghead_Mixinghead{0}_Pressure_Connection{6}_PV_SetV_WarningUpperLimit" : Real = PLC DB604_PV_Mixinghead.Mixinghead[0].Pressure_Connection[6].PV_SetV.WarningUpperLimit AT %DB604.DBD254, 1 s
      on ChangeValue: SetBit("DB704_MH_Value_Write")
   "DB604_PV_Mixinghead_Mixinghead{0}_Pressure_Connection{6}_PV_SetV_AlarmLowerLimit" : Real = PLC DB604_PV_Mixinghead.Mixinghead[0].Pressure_Connection[6].PV_SetV.AlarmLowerLimit AT %DB604.DBD258, 1 s
      on ChangeValue: SetBit("DB704_MH_Value_Write")
   "DB604_PV_Mixinghead_Mixinghead{0}_Pressure_Connection{6}_PV_SetV_AlarmUpperLimit" : Real = PLC DB604_PV_Mixinghead.Mixinghead[0].Pressure_Connection[6].PV_SetV.AlarmUpperLimit AT %DB604.DBD262, 1 s
      on ChangeValue: SetBit("DB704_MH_Value_Write")
   "DB604_PV_Mixinghead_Mixinghead{0}_Pressure_Connection{6}_PV_ActV_Value" : Real = PLC DB604_PV_Mixinghead.Mixinghead[0].Pressure_Connection[6].PV_ActV.Value AT %DB604.DBD266, 1 s
      on ChangeValue: SetBit("DB704_MH_Value_Write")
   "Temp_Name" : WString[20], internal
   "Temp_Actual" : Real, internal
   "Temp_SetValue" : Real, internal
   "Temp_Warning_Upper_Limit" : Real, internal
   "Temp_Warning_Llower_Limit" : Real, internal
   "Temp_Fault_Upper_Limit" : Real, internal
   "Temp_Fault_Lower_Limit" : Real, internal
   "Press_Actual" : Real, internal
   "Press_SetValue" : Real, internal
   "Press_Warning_Upper_Limit" : Real, internal
   "Press_Warning_Lower_Limit" : Real, internal
   "Press_Fault_Upper_Limit" : Real, internal
   "Press_Fault_Lower_Limit" : Real, internal
   "Temp_Control_Screen" : Int, internal
   "Press_Control_Screen" : Int, internal
   "Press_Name" : WString[20], internal
   "DB704_MH_Value_Mixinghead{0}_MH_Connection{1}_WithNozzle" : Bool = PLC DB704_MH_Value.Mixinghead[0].MH_Connection[1].WithNozzle AT %DB704.DBX98.3, 1 s
      on ChangeValue: SetBit("DB704_MH_Value_Write")
   "DB704_MH_Value_Mixinghead{0}_MH_Connection{2}_WithNozzle" : Bool = PLC DB704_MH_Value.Mixinghead[0].MH_Connection[2].WithNozzle AT %DB704.DBX132.3, 1 s
      on ChangeValue: SetBit("DB704_MH_Value_Write")
   "DB704_MH_Value_Mixinghead{0}_MH_Connection{3}_WithNozzle" : Bool = PLC DB704_MH_Value.Mixinghead[0].MH_Connection[3].WithNozzle AT %DB704.DBX166.3, 1 s
      on ChangeValue: SetBit("DB704_MH_Value_Write")
   "DB704_MH_Value_Mixinghead{0}_MH_Connection{4}_WithNozzle" : Bool = PLC DB704_MH_Value.Mixinghead[0].MH_Connection[4].WithNozzle AT %DB704.DBX200.3, 1 s
      on ChangeValue: SetBit("DB704_MH_Value_Write")
   "DB704_MH_Value_Mixinghead{0}_MH_Connection{5}_WithNozzle" : Bool = PLC DB704_MH_Value.Mixinghead[0].MH_Connection[5].WithNozzle AT %DB704.DBX234.3, 1 s
      on ChangeValue: SetBit("DB704_MH_Value_Write")
   "DB704_MH_Value_Mixinghead{0}_DelayTimeNozzlesOff" : S5Time = PLC DB704_MH_Value.Mixinghead[0].DelayTimeNozzlesOff AT %DB704.DBW26, 1 s
      on ChangeValue: SetBit("DB704_MH_Value_Write")
   "DB704_MH_Value_Mixinghead{0}_MH_Connection{6}_WithNozzle" : Bool = PLC DB704_MH_Value.Mixinghead[0].MH_Connection[6].WithNozzle AT %DB704.DBX268.3, 1 s
      on ChangeValue: SetBit("DB704_MH_Value_Write")
   "DB704_MH_Value_MH_Inerting{0}_Inert_Switch_ON_OFF" : Bool = PLC DB704_MH_Value.MH_Inerting[0].Inert_Switch_ON_OFF AT %DB704.DBX4528.7, 1 s
   "DB614_MH_State_MH_Connection{0}_ActFlow{1}" : Real = PLC DB614_MH_State.MH_Connection[0].ActFlow[1] AT %DB614.DBD196, 1 s
   "DB614_MH_State_MH_Connection{0}_ActFlow{2}" : Real = PLC DB614_MH_State.MH_Connection[0].ActFlow[2] AT %DB614.DBD200, 1 s
   "DB614_MH_State_MH_Connection{0}_ActFlow{3}" : Real = PLC DB614_MH_State.MH_Connection[0].ActFlow[3] AT %DB614.DBD204, 1 s
   "DB614_MH_State_MH_Connection{0}_ActFlow{4}" : Real = PLC DB614_MH_State.MH_Connection[0].ActFlow[4] AT %DB614.DBD208, 1 s
   "DB614_MH_State_MH_Connection{0}_ActFlow{5}" : Real = PLC DB614_MH_State.MH_Connection[0].ActFlow[5] AT %DB614.DBD212, 1 s
   "DB614_MH_State_MH_Connection{0}_ActFlow{6}" : Real = PLC DB614_MH_State.MH_Connection[0].ActFlow[6] AT %DB614.DBD216, 1 s
   "DB614_MH_State_InertingMH{0}_Computed_Value" : Real = PLC DB614_MH_State.InertingMH[0].Computed_Value AT %DB614.DBD4302, 1 s
   "DB614_MH_State_InertingMH{0}_Total_Flow_N2_Visu" : Real = PLC DB614_MH_State.InertingMH[0].Total_Flow_N2_Visu AT %DB614.DBD4318, 1 s
   "DB611_Hydraulic_State_MH_Hydraulic{1}_Fault_Exist" : Bool = PLC DB611_Hydraulic_State.MH_Hydraulic[1].Fault_Exist AT %DB611.DBX18.7, 1 s
   "DB614_MH_State_MH_CleaningPiston{0}_Switch_CP_Forward" : Bool = PLC DB614_MH_State.MH_CleaningPiston[0].Switch_CP_Forward AT %DB614.DBX4091.1, 1 s
      on ChangeValue: SetBit("DB614_MH_State_Write")
   "DB614_MH_State_MH_Status{0}_State_HP" : Int = PLC DB614_MH_State.MH_Status[0].State_HP AT %DB614.DBW3922, 1 s
   "DB614_MH_State_MH_Status{0}_State_Service" : Int = PLC DB614_MH_State.MH_Status[0].State_Service AT %DB614.DBW3924, 1 s
   "DB614_MH_State_MH_CleaningPiston{0}_State_CP" : Byte = PLC DB614_MH_State.MH_CleaningPiston[0].State_CP AT %DB614.DBB4094, 1 s
   "DB704_MH_Value_Mixinghead{0}_Corrvalue" : Real = PLC DB704_MH_Value.Mixinghead[0].Corrvalue AT %DB704.DBD62, 1 s
      on ChangeValue: SetBit("DB704_MH_Value_Write")
   "DB704_MH_Value_Mixinghead{0}_Cleaning_Piston_Spare_19" : Bool = PLC DB704_MH_Value.Mixinghead[0].Cleaning_Piston.Spare_19 AT %DB704.DBX56.4, 1 s
      on ChangeValue: SetBit("DB704_MH_Value_Write")
   "DB704_MH_Value_MH_Inerting{0}_with_Purge" : Bool = PLC DB704_MH_Value.MH_Inerting[0].with_Purge AT %DB704.DBX4528.0, 1 s
   "DB704_MH_Value_Mixinghead{0}_Cleaning_Piston_StepCleaningPiston" : Bool = PLC DB704_MH_Value.Mixinghead[0].Cleaning_Piston.StepCleaningPiston AT %DB704.DBX56.2, 1 s
      on ChangeValue: SetBit("DB704_MH_Value_Write")
   "DB704_MH_Value_Mixinghead{0}_Conf_IntWithRobot" : Bool = PLC DB704_MH_Value.Mixinghead[0].Conf_IntWithRobot AT %DB704.DBX10.3, 1 s
      on ChangeValue: SetBit("DB704_MH_Value_Write")
   "DB704_MH_Value_Mixinghead{0}_Conf_IntWithMC" : Bool = PLC DB704_MH_Value.Mixinghead[0].Conf_IntWithMC AT %DB704.DBX10.4, 1 s
      on ChangeValue: SetBit("DB704_MH_Value_Write")
   "DB704_MH_Value_Mixinghead{0}_Conf_IntWithPlantInerface" : Bool = PLC DB704_MH_Value.Mixinghead[0].Conf_IntWithPlantInerface AT %DB704.DBX10.5, 1 s
      on ChangeValue: SetBit("DB704_MH_Value_Write")
   "DB704_MH_Value_Mixinghead{0}_Conf_IntWithCoupler" : Bool = PLC DB704_MH_Value.Mixinghead[0].Conf_IntWithCoupler AT %DB704.DBX10.6, 1 s
      on ChangeValue: SetBit("DB704_MH_Value_Write")
   "DB704_MH_Value_Mixinghead{0}_Conf_IntWithProcessValue" : Bool = PLC DB704_MH_Value.Mixinghead[0].Conf_IntWithProcessValue AT %DB704.DBX10.7, 1 s
      on ChangeValue: SetBit("DB704_MH_Value_Write")
   "DB704_MH_Value_Mixinghead{0}_Conf_IntWithTag" : Bool = PLC DB704_MH_Value.Mixinghead[0].Conf_IntWithTag AT %DB704.DBX11.0, 1 s
      on ChangeValue: SetBit("DB704_MH_Value_Write")
   "DB704_MH_Value_Mixinghead{0}_Conf_MHDigital" : Bool = PLC DB704_MH_Value.Mixinghead[0].Conf_MHDigital AT %DB704.DBX11.1, 1 s
      on ChangeValue: SetBit("DB704_MH_Value_Write")
   "DB704_MH_Value_Mixinghead{0}_Conf_MHControled" : Bool = PLC DB704_MH_Value.Mixinghead[0].Conf_MHControled AT %DB704.DBX11.2, 1 s
      on ChangeValue: SetBit("DB704_MH_Value_Write")
   "DB704_MH_Value_Mixinghead{0}_Conf_MHFibre" : Bool = PLC DB704_MH_Value.Mixinghead[0].Conf_MHFibre AT %DB704.DBX11.3, 1 s
      on ChangeValue: SetBit("DB704_MH_Value_Write")
   "DB704_MH_Value_Mixinghead{0}_Conf_MHSpray" : Bool = PLC DB704_MH_Value.Mixinghead[0].Conf_MHSpray AT %DB704.DBX11.4, 1 s
      on ChangeValue: SetBit("DB704_MH_Value_Write")
   "DB704_MH_Value_Mixinghead{0}_Conf_MHSpecial" : Bool = PLC DB704_MH_Value.Mixinghead[0].Conf_MHSpecial AT %DB704.DBX11.5, 1 s
      on ChangeValue: SetBit("DB704_MH_Value_Write")
   "DB704_MH_Value_MH_Inerting{0}_with_inert_over_MH" : Bool = PLC DB704_MH_Value.MH_Inerting[0].with_inert_over_MH AT %DB704.DBX4528.4, 1 s
      on ChangeValue: SetBit("DB704_MH_Value_Write")
   "DB704_MH_Value_MH_Inerting{0}_with_inert_over_Lance" : Bool = PLC DB704_MH_Value.MH_Inerting[0].with_inert_over_Lance AT %DB704.DBX4528.5, 1 s
      on ChangeValue: SetBit("DB704_MH_Value_Write")
   "DB704_MH_Value_MH_Inerting{0}_with_output_without_N2" : Bool = PLC DB704_MH_Value.MH_Inerting[0].with_output_without_N2 AT %DB704.DBX4528.6, 1 s
      on ChangeValue: SetBit("DB704_MH_Value_Write")
   "DB704_MH_Value_MH_Inerting{0}_Max_Reference_Value_Inert" : Real = PLC DB704_MH_Value.MH_Inerting[0].Max_Reference_Value_Inert AT %DB704.DBD4534, 1 s
      on ChangeValue: SetBit("DB704_MH_Value_Write")
   "DB704_MH_Value_MH_Inerting{0}_Reference_Value_Inert" : Real = PLC DB704_MH_Value.MH_Inerting[0].Reference_Value_Inert AT %DB704.DBD4530, 1 s
   "DB614_MH_State_FaulExist" : Bool = PLC DB614_MH_State.FaulExist AT %DB614.DBX8.5, 1 s
   "DB614_MH_State_MH_Status{0}_FaultExist" : Bool = PLC DB614_MH_State.MH_Status[0].FaultExist AT %DB614.DBX3920.7, 1 s
   "DB123_MH_IO_Signals_MH{0}_IN_MH_Prog_No_MH" : Byte = PLC DB123_MH_IO_Signals.MH[0].IN.MH_Prog_No_MH AT %DB123.DBB2, 1 s
   "DB123_MH_IO_Signals_MH{0}_IN_MH_Manual_Mode" : Bool = PLC DB123_MH_IO_Signals.MH[0].IN.MH_Manual_Mode AT %DB123.DBX0.5, 1 s
      on ChangeValue: "MH_TestshotVisibility"()
   "DB123_MH_IO_Signals_MH{0}_IN_MH_Auto_Mode" : Bool = PLC DB123_MH_IO_Signals.MH[0].IN.MH_Auto_Mode AT %DB123.DBX0.6, 1 s
      on ChangeValue: "MH_TestshotVisibility"()
   "DB614_MH_State_MH_Status{0}_Switch_Testshot_A_ON_OFF" : Bool = PLC DB614_MH_State.MH_Status[0].Switch_Testshot_A_ON_OFF AT %DB614.DBX3921.1, 1 s
      on ChangeValue: SetBit("DB614_MH_State_Write")
   "DB614_MH_State_MH_Status{0}_Switch_Testshot_B_ON_OFF" : Bool = PLC DB614_MH_State.MH_Status[0].Switch_Testshot_B_ON_OFF AT %DB614.DBX3921.2, 1 s
      on ChangeValue: SetBit("DB614_MH_State_Write")
   "DB614_MH_State_MH_Status{0}_State_Testshot_A" : Int = PLC DB614_MH_State.MH_Status[0].State_Testshot_A AT %DB614.DBW3926, 1 s
   "DB614_MH_State_MH_Status{0}_State_Testshot_B" : Int = PLC DB614_MH_State.MH_Status[0].State_Testshot_B AT %DB614.DBW3928, 1 s
   "DB704_MH_Value_Mixinghead{0}_MH_Connection{1}_HP_2Point_Flow" : Bool = PLC DB704_MH_Value.Mixinghead[0].MH_Connection[1].HP_2Point_Flow AT %DB704.DBX98.4, 1 s
   "DB704_MH_Value_Mixinghead{0}_MH_Connection{1}_Red_2Point_Flow" : Bool = PLC DB704_MH_Value.Mixinghead[0].MH_Connection[1].Red_2Point_Flow AT %DB704.DBX98.5, 1 s
   "DB704_MH_Value_Mixinghead{0}_MH_Connection{1}_LP_2Point_Flow" : Bool = PLC DB704_MH_Value.Mixinghead[0].MH_Connection[1].LP_2Point_Flow AT %DB704.DBX98.6, 1 s
   "DB704_MH_Value_Mixinghead{0}_MH_Connection{2}_HP_2Point_Flow" : Bool = PLC DB704_MH_Value.Mixinghead[0].MH_Connection[2].HP_2Point_Flow AT %DB704.DBX132.4, 1 s
   "DB704_MH_Value_Mixinghead{0}_MH_Connection{2}_Red_2Point_Flow" : Bool = PLC DB704_MH_Value.Mixinghead[0].MH_Connection[2].Red_2Point_Flow AT %DB704.DBX132.5, 1 s
   "DB704_MH_Value_Mixinghead{0}_MH_Connection{2}_LP_2Point_Flow" : Bool = PLC DB704_MH_Value.Mixinghead[0].MH_Connection[2].LP_2Point_Flow AT %DB704.DBX132.6, 1 s
   "DB704_MH_Value_Mixinghead{0}_MH_Connection{3}_HP_2Point_Flow" : Bool = PLC DB704_MH_Value.Mixinghead[0].MH_Connection[3].HP_2Point_Flow AT %DB704.DBX166.4, 1 s
   "DB704_MH_Value_Mixinghead{0}_MH_Connection{3}_Red_2Point_Flow" : Bool = PLC DB704_MH_Value.Mixinghead[0].MH_Connection[3].Red_2Point_Flow AT %DB704.DBX166.5, 1 s
   "DB704_MH_Value_Mixinghead{0}_MH_Connection{3}_LP_2Point_Flow" : Bool = PLC DB704_MH_Value.Mixinghead[0].MH_Connection[3].LP_2Point_Flow AT %DB704.DBX166.6, 1 s
   "DB704_MH_Value_Mixinghead{0}_MH_Connection{4}_HP_2Point_Flow" : Bool = PLC DB704_MH_Value.Mixinghead[0].MH_Connection[4].HP_2Point_Flow AT %DB704.DBX200.4, 1 s
   "DB704_MH_Value_Mixinghead{0}_MH_Connection{4}_Red_2Point_Flow" : Bool = PLC DB704_MH_Value.Mixinghead[0].MH_Connection[4].Red_2Point_Flow AT %DB704.DBX200.5, 1 s
   "DB704_MH_Value_Mixinghead{0}_MH_Connection{4}_LP_2Point_Flow" : Bool = PLC DB704_MH_Value.Mixinghead[0].MH_Connection[4].LP_2Point_Flow AT %DB704.DBX200.6, 1 s
   "DB704_MH_Value_Mixinghead{0}_MH_Connection{5}_HP_2Point_Flow" : Bool = PLC DB704_MH_Value.Mixinghead[0].MH_Connection[5].HP_2Point_Flow AT %DB704.DBX234.4, 1 s
   "DB704_MH_Value_Mixinghead{0}_MH_Connection{5}_Red_2Point_Flow" : Bool = PLC DB704_MH_Value.Mixinghead[0].MH_Connection[5].Red_2Point_Flow AT %DB704.DBX234.5, 1 s
   "DB704_MH_Value_Mixinghead{0}_MH_Connection{5}_LP_2Point_Flow" : Bool = PLC DB704_MH_Value.Mixinghead[0].MH_Connection[5].LP_2Point_Flow AT %DB704.DBX234.6, 1 s
   "DB704_MH_Value_Mixinghead{0}_MH_Connection{6}_HP_2Point_Flow" : Bool = PLC DB704_MH_Value.Mixinghead[0].MH_Connection[6].HP_2Point_Flow AT %DB704.DBX268.4, 1 s
   "DB704_MH_Value_Mixinghead{0}_MH_Connection{6}_Red_2Point_Flow" : Bool = PLC DB704_MH_Value.Mixinghead[0].MH_Connection[6].Red_2Point_Flow AT %DB704.DBX268.5, 1 s
   "DB704_MH_Value_Mixinghead{0}_MH_Connection{6}_LP_2Point_Flow" : Bool = PLC DB704_MH_Value.Mixinghead[0].MH_Connection[6].LP_2Point_Flow AT %DB704.DBX268.6, 1 s
   "DB619_State_MPart_Recirculation{1}_Switch_Intervall" : Bool = PLC DB619_State_MPart.Recirculation[1].Switch_Intervall AT %DB619.DBX44.0, 1 s
   "DB619_State_MPart_Recirculation{1}_Switch_Lowpressure" : Bool = PLC DB619_State_MPart.Recirculation[1].Switch_Lowpressure AT %DB619.DBX44.2, 1 s
   "DB619_State_MPart_Recirculation{1}_Switch_Reduced" : Bool = PLC DB619_State_MPart.Recirculation[1].Switch_Reduced AT %DB619.DBX44.3, 1 s
   "DB611_Hydraulic_State_MH_Hydraulic{0}_Fault_Exist" : Bool = PLC DB611_Hydraulic_State.MH_Hydraulic[0].Fault_Exist AT %DB611.DBX10.7, 1 s
   "DB704_MH_Value_Mixinghead{0}_MH_Connection{6}_Pump_No" : Int = PLC DB704_MH_Value.Mixinghead[0].MH_Connection[6].Pump_No AT %DB704.DBW238, 1 s
      on ChangeValue: SetBit("DB704_MH_Value_Write")
   "DB704_MH_Value_Mixinghead{0}_MH_Connection{5}_Pump_No" : Int = PLC DB704_MH_Value.Mixinghead[0].MH_Connection[5].Pump_No AT %DB704.DBW204, 1 s
      on ChangeValue: SetBit("DB704_MH_Value_Write")
   "DB704_MH_Value_Mixinghead{0}_MH_Connection{4}_Pump_No" : Int = PLC DB704_MH_Value.Mixinghead[0].MH_Connection[4].Pump_No AT %DB704.DBW170, 1 s
      on ChangeValue: SetBit("DB704_MH_Value_Write")
   "DB704_MH_Value_Mixinghead{0}_MH_Connection{3}_Pump_No" : Int = PLC DB704_MH_Value.Mixinghead[0].MH_Connection[3].Pump_No AT %DB704.DBW136, 1 s
      on ChangeValue: SetBit("DB704_MH_Value_Write")
   "DB704_MH_Value_Mixinghead{0}_MH_Connection{2}_Pump_No" : Int = PLC DB704_MH_Value.Mixinghead[0].MH_Connection[2].Pump_No AT %DB704.DBW102, 1 s
      on ChangeValue: SetBit("DB704_MH_Value_Write")
   "DB704_MH_Value_Mixinghead{0}_MH_Connection{1}_Pump_No" : Int = PLC DB704_MH_Value.Mixinghead[0].MH_Connection[1].Pump_No AT %DB704.DBW68, 1 s
      on ChangeValue: SetBit("DB704_MH_Value_Write")
   "DB614_MH_State_MH_Connection{0}_Name{1}" : String[20] = PLC DB614_MH_State.MH_Connection[0].Name[1] AT %DB614.DBX10.0, 1 s
   "DB614_MH_State_MH_Connection{0}_Name{2}" : String[20] = PLC DB614_MH_State.MH_Connection[0].Name[2] AT %DB614.DBX32.0, 1 s
   "DB614_MH_State_MH_Connection{0}_Name{3}" : String[20] = PLC DB614_MH_State.MH_Connection[0].Name[3] AT %DB614.DBX54.0, 1 s
   "DB614_MH_State_MH_Connection{0}_Name{4}" : String[20] = PLC DB614_MH_State.MH_Connection[0].Name[4] AT %DB614.DBX76.0, 1 s
   "DB614_MH_State_MH_Connection{0}_Name{5}" : String[20] = PLC DB614_MH_State.MH_Connection[0].Name[5] AT %DB614.DBX98.0, 1 s
   "DB614_MH_State_MH_Connection{0}_Name{6}" : String[20] = PLC DB614_MH_State.MH_Connection[0].Name[6] AT %DB614.DBX120.0, 1 s
   "DB614_MH_State_MH_Connection{0}_colour{1}" : Byte = PLC DB614_MH_State.MH_Connection[0].colour[1] AT %DB614.DBB142, 1 s
   "DB614_MH_State_MH_Connection{0}_colour{2}" : Byte = PLC DB614_MH_State.MH_Connection[0].colour[2] AT %DB614.DBB143, 1 s
   "DB614_MH_State_MH_Connection{0}_colour{3}" : Byte = PLC DB614_MH_State.MH_Connection[0].colour[3] AT %DB614.DBB144, 1 s
   "DB614_MH_State_MH_Connection{0}_colour{4}" : Byte = PLC DB_MouldEditor_HMI.uData.arShotSet[5].Flow[4] AT %DB614.DBB145, 1 s
   "DB614_MH_State_MH_Connection{0}_colour{5}" : Byte = PLC DB614_MH_State.MH_Connection[0].colour[5] AT %DB614.DBB146, 1 s
   "DB614_MH_State_MH_Connection{0}_colour{6}" : Byte = PLC DB614_MH_State.MH_Connection[0].colour[6] AT %DB614.DBB147, 1 s
   "DB123_MH_IO_Signals_MH{0}_IN_MH_Opentime" : Real = PLC DB123_MH_IO_Signals.MH[0].IN.MH_Opentime AT %DB123.DBD8, 1 s
   "DB123_MH_IO_Signals_MH{0}_IN_MH_Closingtime" : Real = PLC DB123_MH_IO_Signals.MH[0].IN.MH_Closingtime AT %DB123.DBD12, 1 s
   "DB704_MH_Value_Mixinghead{0}_Cleaning_Piston_IntervalCounts" : Int = PLC DB704_MH_Value.Mixinghead[0].Cleaning_Piston.IntervalCounts AT %DB704.DBW50, 1 s
      on ChangeValue: SetBit("DB704_MH_Value_Write")
   "DB704_MH_Value_Mixinghead{0}_Cleaning_Piston_IntervalRestTimeBack" : S5Time = PLC DB704_MH_Value.Mixinghead[0].Cleaning_Piston.IntervalRestTimeBack AT %DB704.DBW52, 1 s
      on ChangeValue: SetBit("DB704_MH_Value_Write")
   "DB704_MH_Value_Mixinghead{0}_Cleaning_Piston_IntervalRestTimeFront" : S5Time = PLC DB704_MH_Value.Mixinghead[0].Cleaning_Piston.IntervalRestTimeFront AT %DB704.DBW54, 1 s
      on ChangeValue: SetBit("DB704_MH_Value_Write")
   "DB619_State_MPart_SWU{1}_ActualSWU" : Int = PLC DB619_State_MPart.SWU[1].ActualSWU AT %DB619.DBW124, 1 s

